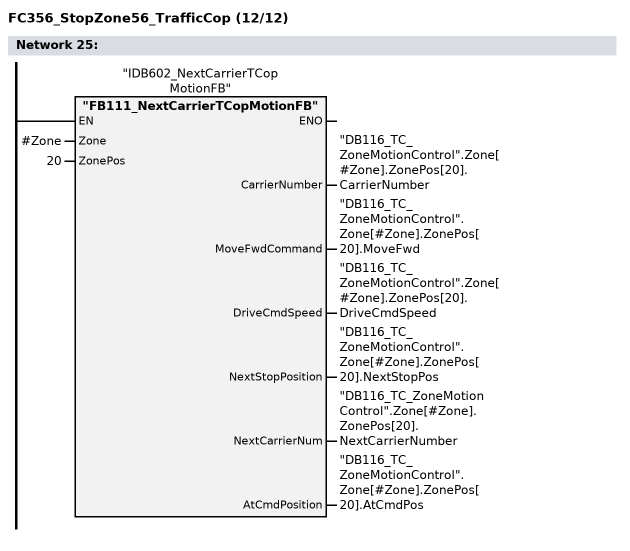
   RUNG wire#powerrail
      "IDB602_NextCarrierTCopMotionFB"(Zone := #Zone, ZonePos := 20, CarrierNumber => "DB116_TC_ZoneMotionControl".Zone[#Zone].ZonePos[20].CarrierNumber, MoveFwdCommand => "DB116_TC_ZoneMotionControl".Zone[#Zone].ZonePos[20].MoveFwd, DriveCmdSpeed => "DB116_TC_ZoneMotionControl".Zone[#Zone].ZonePos[20].DriveCmdSpeed, NextStopPosition => "DB116_TC_ZoneMotionControl".Zone[#Zone].ZonePos[20].NextStopPos, NextCarrierNum => "DB116_TC_ZoneMotionControl".Zone[#Zone].ZonePos[20].NextCarrierNumber, AtCmdPosition => "DB116_TC_ZoneMotionControl".Zone[#Zone].ZonePos[20].AtCmdPos)
   END_RUNG
   // the same network as SCL:
   "IDB602_NextCarrierTCopMotionFB"(Zone := #Zone,   // "FB111_NextCarrierTCopMotionFB"
                           ZonePos := 20,
                           CarrierNumber => "DB116_TC_ZoneMotionControl".Zone[#Zone].ZonePos[20].CarrierNumber,
                           MoveFwdCommand => "DB116_TC_ZoneMotionControl".Zone[#Zone].ZonePos[20].MoveFwd,
                           DriveCmdSpeed => "DB116_TC_ZoneMotionControl".Zone[#Zone].ZonePos[20].DriveCmdSpeed,
                           NextStopPosition => "DB116_TC_ZoneMotionControl".Zone[#Zone].ZonePos[20].NextStopPos,
                           NextCarrierNum => "DB116_TC_ZoneMotionControl".Zone[#Zone].ZonePos[20].NextCarrierNumber,
                           AtCmdPosition => "DB116_TC_ZoneMotionControl".Zone[#Zone].ZonePos[20].AtCmdPos);
END_REGION
END_FUNCTION

FUNCTION "FC357_StopZone57_TrafficCop" : Void   // FC357, LAD
{ S7_Optimized_Access := 'FALSE' }
VERSION : 0.1
   VAR_INPUT
      Zone : Int;
   END_VAR
   VAR_TEMP
      TrafficCopCarrier : Int;
      CarrierMotionZn : Array[0..40] of "UDT_ZoneCarrierStatus";
   END_VAR
BEGIN

REGION Network 1
   // **********************************************************************************************************************
   // 
   // Zone Function Block.  Static setup of all Zone Parameters.  Traffic Cop Setup Logic - Handles all motion and carrier movement logic based on interdependence of Each Carrier in Zone # Passed from Main program Call in OB1 
   // 
   // **********************************************************************************************************************
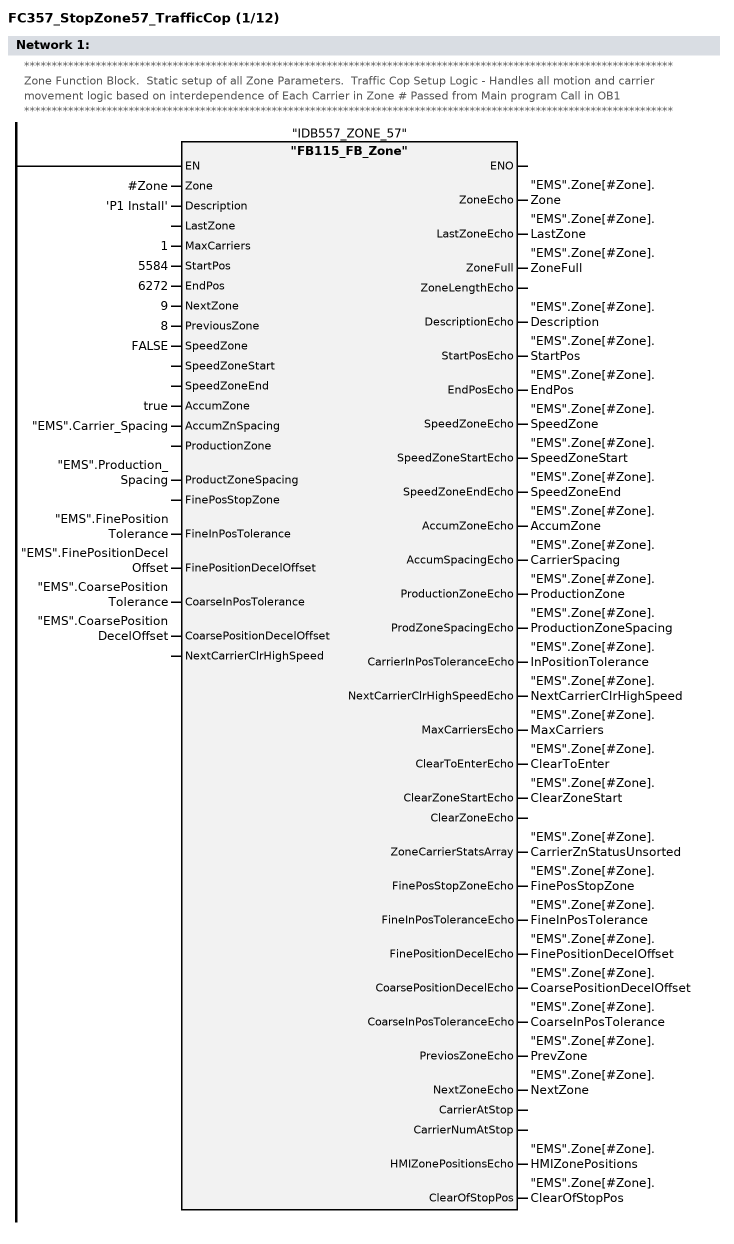
   RUNG wire#powerrail
      "IDB557_ZONE_57"(Zone := #Zone, Description := 'P1 Install', LastZone :=, MaxCarriers := 1, StartPos := 5584, EndPos := 6272, NextZone := 9, PreviousZone := 8, SpeedZone := FALSE, SpeedZoneStart :=, SpeedZoneEnd :=, AccumZone := true, AccumZnSpacing := "EMS".Carrier_Spacing, ProductionZone :=, ProductZoneSpacing := "EMS".Production_Spacing, FinePosStopZone :=, FineInPosTolerance := "EMS".FinePositionTolerance, FinePositionDecelOffset := "EMS".FinePositionDecelOffset, CoarseInPosTolerance := "EMS".CoarsePositionTolerance, CoarsePositionDecelOffset := "EMS".CoarsePositionDecelOffset, NextCarrierClrHighSpeed :=, ZoneEcho => "EMS".Zone[#Zone].Zone, LastZoneEcho => "EMS".Zone[#Zone].LastZone, ZoneFull => "EMS".Zone[#Zone].ZoneFull, ZoneLengthEcho =>, DescriptionEcho => "EMS".Zone[#Zone].Description, StartPosEcho => "EMS".Zone[#Zone].StartPos, EndPosEcho => "EMS".Zone[#Zone].EndPos, SpeedZoneEcho => "EMS".Zone[#Zone].SpeedZone, SpeedZoneStartEcho => "EMS".Zone[#Zone].SpeedZoneStart, SpeedZoneEndEcho => "EMS".Zone[#Zone].SpeedZoneEnd, AccumZoneEcho => "EMS".Zone[#Zone].AccumZone, AccumSpacingEcho => "EMS".Zone[#Zone].CarrierSpacing, ProductionZoneEcho => "EMS".Zone[#Zone].ProductionZone, ProdZoneSpacingEcho => "EMS".Zone[#Zone].ProductionZoneSpacing, CarrierInPosToleranceEcho => "EMS".Zone[#Zone].InPositionTolerance, NextCarrierClrHighSpeedEcho => "EMS".Zone[#Zone].NextCarrierClrHighSpeed, MaxCarriersEcho => "EMS".Zone[#Zone].MaxCarriers, ClearToEnterEcho => "EMS".Zone[#Zone].ClearToEnter, ClearZoneStartEcho => "EMS".Zone[#Zone].ClearZoneStart, ClearZoneEcho =>, ZoneCarrierStatsArray => "EMS".Zone[#Zone].CarrierZnStatusUnsorted, FinePosStopZoneEcho => "EMS".Zone[#Zone].FinePosStopZone, FineInPosToleranceEcho => "EMS".Zone[#Zone].FineInPosTolerance, FinePositionDecelEcho => "EMS".Zone[#Zone].FinePositionDecelOffset, CoarsePositionDecelEcho => "EMS".Zone[#Zone].CoarsePositionDecelOffset, CoarseInPosToleranceEcho => "EMS".Zone[#Zone].CoarseInPosTolerance, PreviosZoneEcho => "EMS".Zone[#Zone].PrevZone, NextZoneEcho => "EMS".Zone[#Zone].NextZone, CarrierAtStop =>, CarrierNumAtStop =>, HMIZonePositionsEcho => "EMS".Zone[#Zone].HMIZonePositions, ClearOfStopPos => "EMS".Zone[#Zone].ClearOfStopPos)
   END_RUNG
   // the same network as SCL:
   "IDB557_ZONE_57"(Zone := #Zone,   // "FB115_FB_Zone"
                    Description := 'P1 Install',
                    MaxCarriers := 1,
                    StartPos := 5584,
                    EndPos := 6272,
                    NextZone := 9,
                    PreviousZone := 8,
                    SpeedZone := FALSE,
                    AccumZone := true,
                    AccumZnSpacing := "EMS".Carrier_Spacing,
                    ProductZoneSpacing := "EMS".Production_Spacing,
                    FineInPosTolerance := "EMS".FinePositionTolerance,
                    FinePositionDecelOffset := "EMS".FinePositionDecelOffset,
                    CoarseInPosTolerance := "EMS".CoarsePositionTolerance,
                    CoarsePositionDecelOffset := "EMS".CoarsePositionDecelOffset,
                    ZoneEcho => "EMS".Zone[#Zone].Zone,
                    LastZoneEcho => "EMS".Zone[#Zone].LastZone,
                    ZoneFull => "EMS".Zone[#Zone].ZoneFull,
                    DescriptionEcho => "EMS".Zone[#Zone].Description,
                    StartPosEcho => "EMS".Zone[#Zone].StartPos,
                    EndPosEcho => "EMS".Zone[#Zone].EndPos,
                    SpeedZoneEcho => "EMS".Zone[#Zone].SpeedZone,
                    SpeedZoneStartEcho => "EMS".Zone[#Zone].SpeedZoneStart,
                    SpeedZoneEndEcho => "EMS".Zone[#Zone].SpeedZoneEnd,
                    AccumZoneEcho => "EMS".Zone[#Zone].AccumZone,
                    AccumSpacingEcho => "EMS".Zone[#Zone].CarrierSpacing,
                    ProductionZoneEcho => "EMS".Zone[#Zone].ProductionZone,
                    ProdZoneSpacingEcho => "EMS".Zone[#Zone].ProductionZoneSpacing,
                    CarrierInPosToleranceEcho => "EMS".Zone[#Zone].InPositionTolerance,
                    NextCarrierClrHighSpeedEcho => "EMS".Zone[#Zone].NextCarrierClrHighSpeed,
                    MaxCarriersEcho => "EMS".Zone[#Zone].MaxCarriers,
                    ClearToEnterEcho => "EMS".Zone[#Zone].ClearToEnter,
                    ClearZoneStartEcho => "EMS".Zone[#Zone].ClearZoneStart,
                    ZoneCarrierStatsArray => "EMS".Zone[#Zone].CarrierZnStatusUnsorted,
                    FinePosStopZoneEcho => "EMS".Zone[#Zone].FinePosStopZone,
                    FineInPosToleranceEcho => "EMS".Zone[#Zone].FineInPosTolerance,
                    FinePositionDecelEcho => "EMS".Zone[#Zone].FinePositionDecelOffset,
                    CoarsePositionDecelEcho => "EMS".Zone[#Zone].CoarsePositionDecelOffset,
                    CoarseInPosToleranceEcho => "EMS".Zone[#Zone].CoarseInPosTolerance,
                    PreviosZoneEcho => "EMS".Zone[#Zone].PrevZone,
                    NextZoneEcho => "EMS".Zone[#Zone].NextZone,
                    HMIZonePositionsEcho => "EMS".Zone[#Zone].HMIZonePositions,
                    ClearOfStopPos => "EMS".Zone[#Zone].ClearOfStopPos);
END_REGION

REGION Network 2
   // *********************************************************************************************************************
   // Carrier Sort Function FC202 - Sorts Carriers in Called Zone to place in correct sequence within  zone. Zones are divided into position based on MaxCarriers allowed in zone as set in the zone setup function block. 
   // 
   // **********************************************************************************************************************
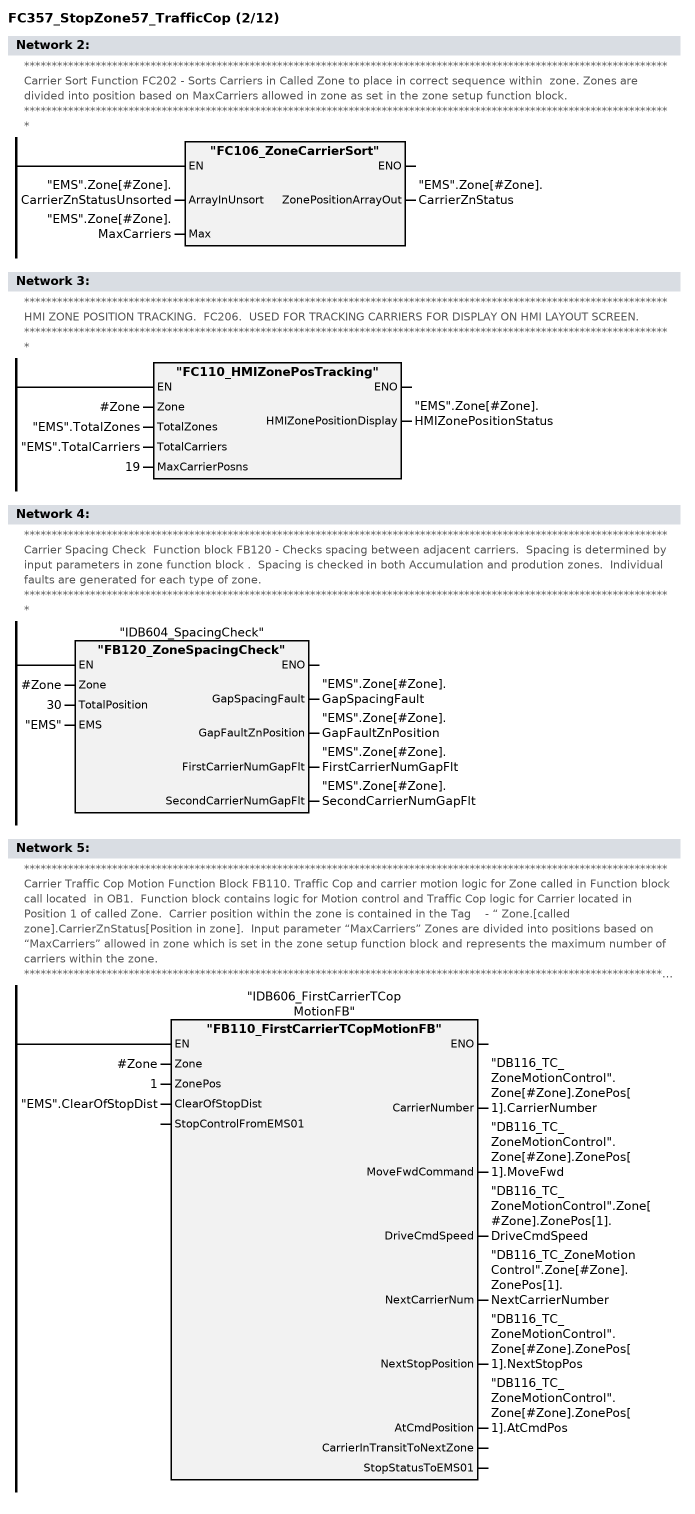
   RUNG wire#powerrail
      "FC106_ZoneCarrierSort"(ArrayInUnsort := "EMS".Zone[#Zone].CarrierZnStatusUnsorted, Max := "EMS".Zone[#Zone].MaxCarriers, ZonePositionArrayOut => "EMS".Zone[#Zone].CarrierZnStatus)
   END_RUNG
   // the same network as SCL:
   "FC106_ZoneCarrierSort"(ArrayInUnsort := "EMS".Zone[#Zone].CarrierZnStatusUnsorted,
                           Max := "EMS".Zone[#Zone].MaxCarriers,
                           ZonePositionArrayOut => "EMS".Zone[#Zone].CarrierZnStatus);
END_REGION

REGION Network 3
   // *********************************************************************************************************************
   // HMI ZONE POSITION TRACKING.  FC206.  USED FOR TRACKING CARRIERS FOR DISPLAY ON HMI LAYOUT SCREEN. 
   // **********************************************************************************************************************
   RUNG wire#powerrail
      "FC110_HMIZonePosTracking"(Zone := #Zone, TotalZones := "EMS".TotalZones, TotalCarriers := "EMS".TotalCarriers, MaxCarrierPosns := 19, HMIZonePositionDisplay => "EMS".Zone[#Zone].HMIZonePositionStatus)
   END_RUNG
   // the same network as SCL:
   "FC110_HMIZonePosTracking"(Zone := #Zone,
                           TotalZones := "EMS".TotalZones,
                           TotalCarriers := "EMS".TotalCarriers,
                           MaxCarrierPosns := 19,
                           HMIZonePositionDisplay => "EMS".Zone[#Zone].HMIZonePositionStatus);
END_REGION

REGION Network 4
   // *********************************************************************************************************************
   // 
   // Carrier Spacing Check  Function block FB120 - Checks spacing between adjacent carriers.  Spacing is determined by input parameters in zone function block .  Spacing is checked in both Accumulation and prodution zones.  Individual faults are generated for each type of zone.
   // 
   // **********************************************************************************************************************
   RUNG wire#powerrail
      "IDB604_SpacingCheck"(Zone := #Zone, TotalPosition := 30, EMS := "EMS", GapSpacingFault => "EMS".Zone[#Zone].GapSpacingFault, GapFaultZnPosition => "EMS".Zone[#Zone].GapFaultZnPosition, FirstCarrierNumGapFlt => "EMS".Zone[#Zone].FirstCarrierNumGapFlt, SecondCarrierNumGapFlt => "EMS".Zone[#Zone].SecondCarrierNumGapFlt)
   END_RUNG
   // the same network as SCL:
   "IDB604_SpacingCheck"(Zone := #Zone,   // "FB120_ZoneSpacingCheck"
                         TotalPosition := 30,
                         EMS := "EMS",
                         GapSpacingFault => "EMS".Zone[#Zone].GapSpacingFault,
                         GapFaultZnPosition => "EMS".Zone[#Zone].GapFaultZnPosition,
                         FirstCarrierNumGapFlt => "EMS".Zone[#Zone].FirstCarrierNumGapFlt,
                         SecondCarrierNumGapFlt => "EMS".Zone[#Zone].SecondCarrierNumGapFlt);
END_REGION

REGION Network 5
   // *********************************************************************************************************************
   // 
   // Carrier Traffic Cop Motion Function Block FB110. Traffic Cop and carrier motion logic for Zone called in Function block call located  in OB1.  Function block contains logic for Motion control and Traffic Cop logic for Carrier located in Position 1 of called Zone.  Carrier position within the zone is contained in the Tag    - “ Zone.[called zone].CarrierZnStatus[Position in zone].  Input parameter “MaxCarriers” Zones are divided into positions based on “MaxCarriers” allowed in zone which is set in the zone setup function block and represents the maximum number of carriers within the zone. 
   // 
   // **********************************************************************************************************************
   RUNG wire#powerrail
      "IDB606_FirstCarrierTCopMotionFB"(Zone := #Zone, ZonePos := 1, ClearOfStopDist := "EMS".ClearOfStopDist, CarrierNumber => "DB116_TC_ZoneMotionControl".Zone[#Zone].ZonePos[1].CarrierNumber, MoveFwdCommand => "DB116_TC_ZoneMotionControl".Zone[#Zone].ZonePos[1].MoveFwd, DriveCmdSpeed => "DB116_TC_ZoneMotionControl".Zone[#Zone].ZonePos[1].DriveCmdSpeed, NextCarrierNum => "DB116_TC_ZoneMotionControl".Zone[#Zone].ZonePos[1].NextCarrierNumber, NextStopPosition => "DB116_TC_ZoneMotionControl".Zone[#Zone].ZonePos[1].NextStopPos, AtCmdPosition => "DB116_TC_ZoneMotionControl".Zone[#Zone].ZonePos[1].AtCmdPos, CarrierInTransitToNextZone =>, StopControlFromEMS01 :=, StopStatusToEMS01 =>)
   END_RUNG
   // the same network as SCL:
   "IDB606_FirstCarrierTCopMotionFB"(Zone := #Zone,   // "FB110_FirstCarrierTCopMotionFB"
                           ZonePos := 1,
                           ClearOfStopDist := "EMS".ClearOfStopDist,
                           CarrierNumber => "DB116_TC_ZoneMotionControl".Zone[#Zone].ZonePos[1].CarrierNumber,
                           MoveFwdCommand => "DB116_TC_ZoneMotionControl".Zone[#Zone].ZonePos[1].MoveFwd,
                           DriveCmdSpeed => "DB116_TC_ZoneMotionControl".Zone[#Zone].ZonePos[1].DriveCmdSpeed,
                           NextCarrierNum => "DB116_TC_ZoneMotionControl".Zone[#Zone].ZonePos[1].NextCarrierNumber,
                           NextStopPosition => "DB116_TC_ZoneMotionControl".Zone[#Zone].ZonePos[1].NextStopPos,
                           AtCmdPosition => "DB116_TC_ZoneMotionControl".Zone[#Zone].ZonePos[1].AtCmdPos);
END_REGION

REGION Network 6
   // *********************************************************************************************************************
   // 
   // Carrier Traffic Cop Motion Function Block FB111. Traffic Cop and carrier motion logic for Zone called in Function block call located  in OB1.  Function block contains logic for Motion control and Traffic Cop logic for Carrier located in Position 2 of called Zone.  Carrier position within the zone is contained in the Tag    - “ Zone.[called zone].CarrierZnStatus[Position in zone].  Input parameter “MaxCarriers” Zones are divided into positions based on “MaxCarriers” allowed in zone which is set in the zone setup function block and represents the maximum number of carriers within the zone. 
   // 
   // **********************************************************************************************************************
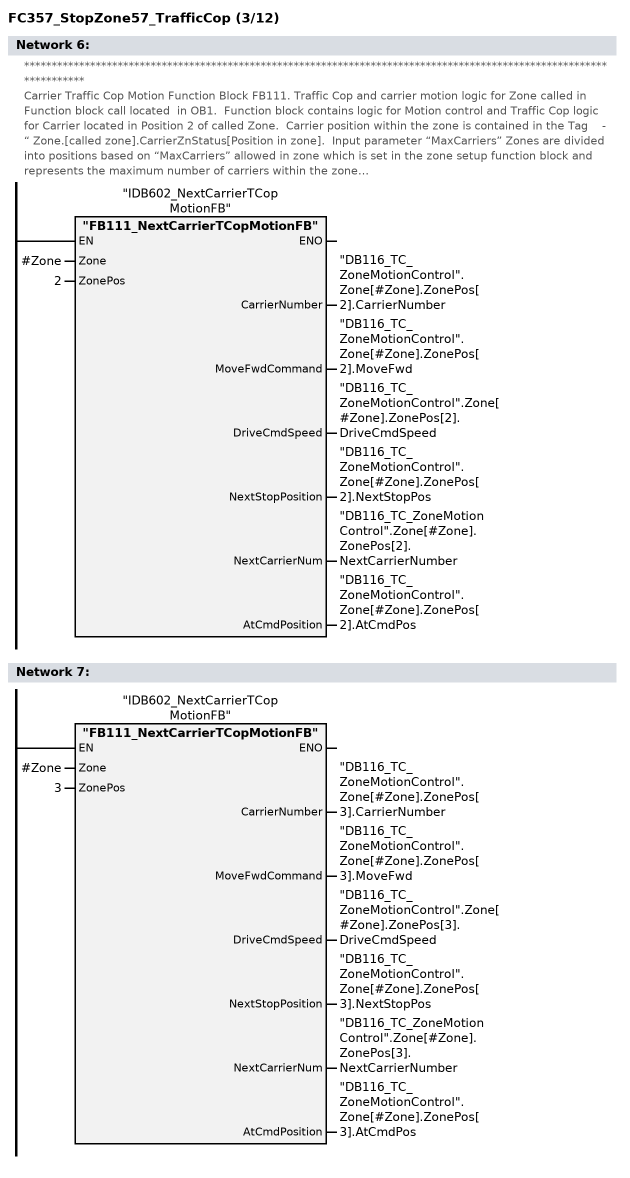
   RUNG wire#powerrail
      "IDB602_NextCarrierTCopMotionFB"(Zone := #Zone, ZonePos := 2, CarrierNumber => "DB116_TC_ZoneMotionControl".Zone[#Zone].ZonePos[2].CarrierNumber, MoveFwdCommand => "DB116_TC_ZoneMotionControl".Zone[#Zone].ZonePos[2].MoveFwd, DriveCmdSpeed => "DB116_TC_ZoneMotionControl".Zone[#Zone].ZonePos[2].DriveCmdSpeed, NextStopPosition => "DB116_TC_ZoneMotionControl".Zone[#Zone].ZonePos[2].NextStopPos, NextCarrierNum => "DB116_TC_ZoneMotionControl".Zone[#Zone].ZonePos[2].NextCarrierNumber, AtCmdPosition => "DB116_TC_ZoneMotionControl".Zone[#Zone].ZonePos[2].AtCmdPos)
   END_RUNG
   // the same network as SCL:
   "IDB602_NextCarrierTCopMotionFB"(Zone := #Zone,   // "FB111_NextCarrierTCopMotionFB"
                           ZonePos := 2,
                           CarrierNumber => "DB116_TC_ZoneMotionControl".Zone[#Zone].ZonePos[2].CarrierNumber,
                           MoveFwdCommand => "DB116_TC_ZoneMotionControl".Zone[#Zone].ZonePos[2].MoveFwd,
                           DriveCmdSpeed => "DB116_TC_ZoneMotionControl".Zone[#Zone].ZonePos[2].DriveCmdSpeed,
                           NextStopPosition => "DB116_TC_ZoneMotionControl".Zone[#Zone].ZonePos[2].NextStopPos,
                           NextCarrierNum => "DB116_TC_ZoneMotionControl".Zone[#Zone].ZonePos[2].NextCarrierNumber,
                           AtCmdPosition => "DB116_TC_ZoneMotionControl".Zone[#Zone].ZonePos[2].AtCmdPos);
END_REGION

REGION Network 7
   RUNG wire#powerrail
      "IDB602_NextCarrierTCopMotionFB"(Zone := #Zone, ZonePos := 3, CarrierNumber => "DB116_TC_ZoneMotionControl".Zone[#Zone].ZonePos[3].CarrierNumber, MoveFwdCommand => "DB116_TC_ZoneMotionControl".Zone[#Zone].ZonePos[3].MoveFwd, DriveCmdSpeed => "DB116_TC_ZoneMotionControl".Zone[#Zone].ZonePos[3].DriveCmdSpeed, NextStopPosition => "DB116_TC_ZoneMotionControl".Zone[#Zone].ZonePos[3].NextStopPos, NextCarrierNum => "DB116_TC_ZoneMotionControl".Zone[#Zone].ZonePos[3].NextCarrierNumber, AtCmdPosition => "DB116_TC_ZoneMotionControl".Zone[#Zone].ZonePos[3].AtCmdPos)
   END_RUNG
   // the same network as SCL:
   "IDB602_NextCarrierTCopMotionFB"(Zone := #Zone,   // "FB111_NextCarrierTCopMotionFB"
                           ZonePos := 3,
                           CarrierNumber => "DB116_TC_ZoneMotionControl".Zone[#Zone].ZonePos[3].CarrierNumber,
                           MoveFwdCommand => "DB116_TC_ZoneMotionControl".Zone[#Zone].ZonePos[3].MoveFwd,
                           DriveCmdSpeed => "DB116_TC_ZoneMotionControl".Zone[#Zone].ZonePos[3].DriveCmdSpeed,
                           NextStopPosition => "DB116_TC_ZoneMotionControl".Zone[#Zone].ZonePos[3].NextStopPos,
                           NextCarrierNum => "DB116_TC_ZoneMotionControl".Zone[#Zone].ZonePos[3].NextCarrierNumber,
                           AtCmdPosition => "DB116_TC_ZoneMotionControl".Zone[#Zone].ZonePos[3].AtCmdPos);
END_REGION

REGION Network 8
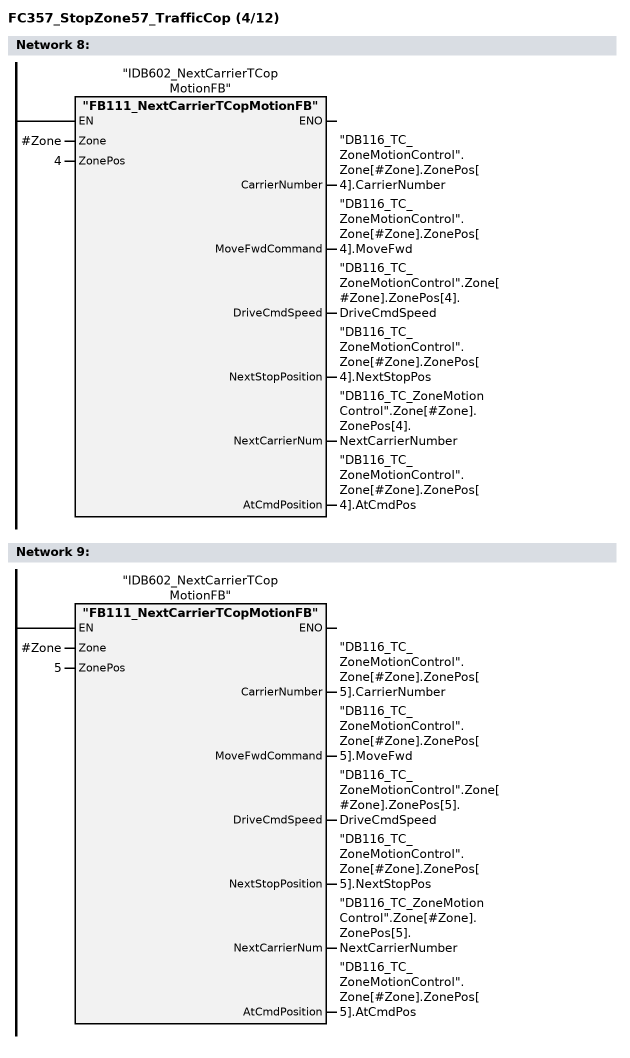
   RUNG wire#powerrail
      "IDB602_NextCarrierTCopMotionFB"(Zone := #Zone, ZonePos := 4, CarrierNumber => "DB116_TC_ZoneMotionControl".Zone[#Zone].ZonePos[4].CarrierNumber, MoveFwdCommand => "DB116_TC_ZoneMotionControl".Zone[#Zone].ZonePos[4].MoveFwd, DriveCmdSpeed => "DB116_TC_ZoneMotionControl".Zone[#Zone].ZonePos[4].DriveCmdSpeed, NextStopPosition => "DB116_TC_ZoneMotionControl".Zone[#Zone].ZonePos[4].NextStopPos, NextCarrierNum => "DB116_TC_ZoneMotionControl".Zone[#Zone].ZonePos[4].NextCarrierNumber, AtCmdPosition => "DB116_TC_ZoneMotionControl".Zone[#Zone].ZonePos[4].AtCmdPos)
   END_RUNG
   // the same network as SCL:
   "IDB602_NextCarrierTCopMotionFB"(Zone := #Zone,   // "FB111_NextCarrierTCopMotionFB"
                           ZonePos := 4,
                           CarrierNumber => "DB116_TC_ZoneMotionControl".Zone[#Zone].ZonePos[4].CarrierNumber,
                           MoveFwdCommand => "DB116_TC_ZoneMotionControl".Zone[#Zone].ZonePos[4].MoveFwd,
                           DriveCmdSpeed => "DB116_TC_ZoneMotionControl".Zone[#Zone].ZonePos[4].DriveCmdSpeed,
                           NextStopPosition => "DB116_TC_ZoneMotionControl".Zone[#Zone].ZonePos[4].NextStopPos,
                           NextCarrierNum => "DB116_TC_ZoneMotionControl".Zone[#Zone].ZonePos[4].NextCarrierNumber,
                           AtCmdPosition => "DB116_TC_ZoneMotionControl".Zone[#Zone].ZonePos[4].AtCmdPos);
END_REGION

REGION Network 9
   RUNG wire#powerrail
      "IDB602_NextCarrierTCopMotionFB"(Zone := #Zone, ZonePos := 5, CarrierNumber => "DB116_TC_ZoneMotionControl".Zone[#Zone].ZonePos[5].CarrierNumber, MoveFwdCommand => "DB116_TC_ZoneMotionControl".Zone[#Zone].ZonePos[5].MoveFwd, DriveCmdSpeed => "DB116_TC_ZoneMotionControl".Zone[#Zone].ZonePos[5].DriveCmdSpeed, NextStopPosition => "DB116_TC_ZoneMotionControl".Zone[#Zone].ZonePos[5].NextStopPos, NextCarrierNum => "DB116_TC_ZoneMotionControl".Zone[#Zone].ZonePos[5].NextCarrierNumber, AtCmdPosition => "DB116_TC_ZoneMotionControl".Zone[#Zone].ZonePos[5].AtCmdPos)
   END_RUNG
   // the same network as SCL:
   "IDB602_NextCarrierTCopMotionFB"(Zone := #Zone,   // "FB111_NextCarrierTCopMotionFB"
                           ZonePos := 5,
                           CarrierNumber => "DB116_TC_ZoneMotionControl".Zone[#Zone].ZonePos[5].CarrierNumber,
                           MoveFwdCommand => "DB116_TC_ZoneMotionControl".Zone[#Zone].ZonePos[5].MoveFwd,
                           DriveCmdSpeed => "DB116_TC_ZoneMotionControl".Zone[#Zone].ZonePos[5].DriveCmdSpeed,
                           NextStopPosition => "DB116_TC_ZoneMotionControl".Zone[#Zone].ZonePos[5].NextStopPos,
                           NextCarrierNum => "DB116_TC_ZoneMotionControl".Zone[#Zone].ZonePos[5].NextCarrierNumber,
                           AtCmdPosition => "DB116_TC_ZoneMotionControl".Zone[#Zone].ZonePos[5].AtCmdPos);
END_REGION

REGION Network 10
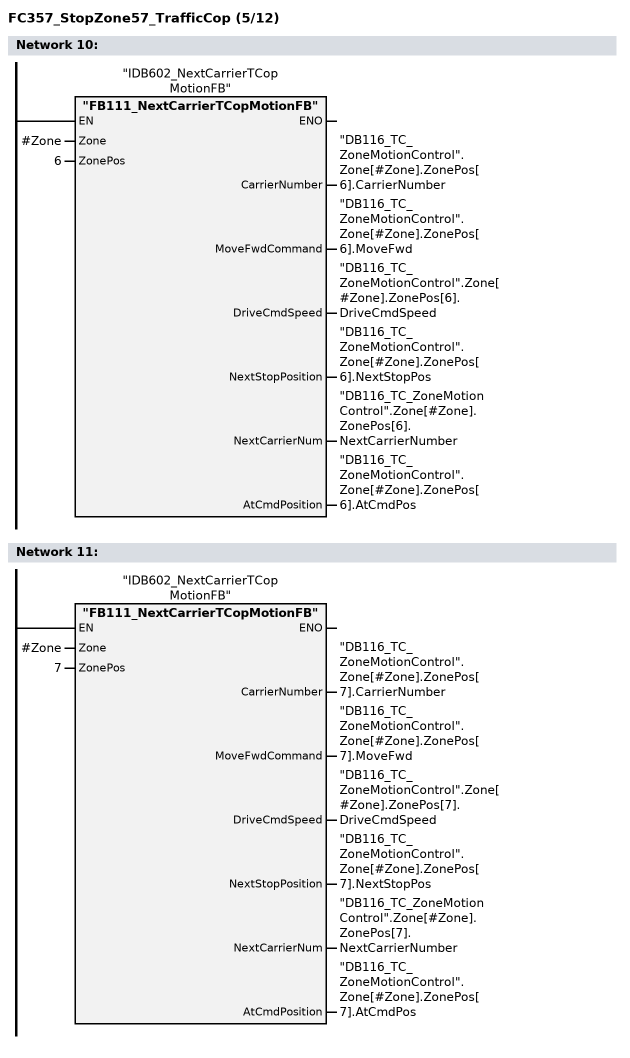
   RUNG wire#powerrail
      "IDB602_NextCarrierTCopMotionFB"(Zone := #Zone, ZonePos := 6, CarrierNumber => "DB116_TC_ZoneMotionControl".Zone[#Zone].ZonePos[6].CarrierNumber, MoveFwdCommand => "DB116_TC_ZoneMotionControl".Zone[#Zone].ZonePos[6].MoveFwd, DriveCmdSpeed => "DB116_TC_ZoneMotionControl".Zone[#Zone].ZonePos[6].DriveCmdSpeed, NextStopPosition => "DB116_TC_ZoneMotionControl".Zone[#Zone].ZonePos[6].NextStopPos, NextCarrierNum => "DB116_TC_ZoneMotionControl".Zone[#Zone].ZonePos[6].NextCarrierNumber, AtCmdPosition => "DB116_TC_ZoneMotionControl".Zone[#Zone].ZonePos[6].AtCmdPos)
   END_RUNG
   // the same network as SCL:
   "IDB602_NextCarrierTCopMotionFB"(Zone := #Zone,   // "FB111_NextCarrierTCopMotionFB"
                           ZonePos := 6,
                           CarrierNumber => "DB116_TC_ZoneMotionControl".Zone[#Zone].ZonePos[6].CarrierNumber,
                           MoveFwdCommand => "DB116_TC_ZoneMotionControl".Zone[#Zone].ZonePos[6].MoveFwd,
                           DriveCmdSpeed => "DB116_TC_ZoneMotionControl".Zone[#Zone].ZonePos[6].DriveCmdSpeed,
                           NextStopPosition => "DB116_TC_ZoneMotionControl".Zone[#Zone].ZonePos[6].NextStopPos,
                           NextCarrierNum => "DB116_TC_ZoneMotionControl".Zone[#Zone].ZonePos[6].NextCarrierNumber,
                           AtCmdPosition => "DB116_TC_ZoneMotionControl".Zone[#Zone].ZonePos[6].AtCmdPos);
END_REGION

REGION Network 11
   RUNG wire#powerrail
      "IDB602_NextCarrierTCopMotionFB"(Zone := #Zone, ZonePos := 7, CarrierNumber => "DB116_TC_ZoneMotionControl".Zone[#Zone].ZonePos[7].CarrierNumber, MoveFwdCommand => "DB116_TC_ZoneMotionControl".Zone[#Zone].ZonePos[7].MoveFwd, DriveCmdSpeed => "DB116_TC_ZoneMotionControl".Zone[#Zone].ZonePos[7].DriveCmdSpeed, NextStopPosition => "DB116_TC_ZoneMotionControl".Zone[#Zone].ZonePos[7].NextStopPos, NextCarrierNum => "DB116_TC_ZoneMotionControl".Zone[#Zone].ZonePos[7].NextCarrierNumber, AtCmdPosition => "DB116_TC_ZoneMotionControl".Zone[#Zone].ZonePos[7].AtCmdPos)
   END_RUNG
   // the same network as SCL:
   "IDB602_NextCarrierTCopMotionFB"(Zone := #Zone,   // "FB111_NextCarrierTCopMotionFB"
                           ZonePos := 7,
                           CarrierNumber => "DB116_TC_ZoneMotionControl".Zone[#Zone].ZonePos[7].CarrierNumber,
                           MoveFwdCommand => "DB116_TC_ZoneMotionControl".Zone[#Zone].ZonePos[7].MoveFwd,
                           DriveCmdSpeed => "DB116_TC_ZoneMotionControl".Zone[#Zone].ZonePos[7].DriveCmdSpeed,
                           NextStopPosition => "DB116_TC_ZoneMotionControl".Zone[#Zone].ZonePos[7].NextStopPos,
                           NextCarrierNum => "DB116_TC_ZoneMotionControl".Zone[#Zone].ZonePos[7].NextCarrierNumber,
                           AtCmdPosition => "DB116_TC_ZoneMotionControl".Zone[#Zone].ZonePos[7].AtCmdPos);
END_REGION

REGION Network 12
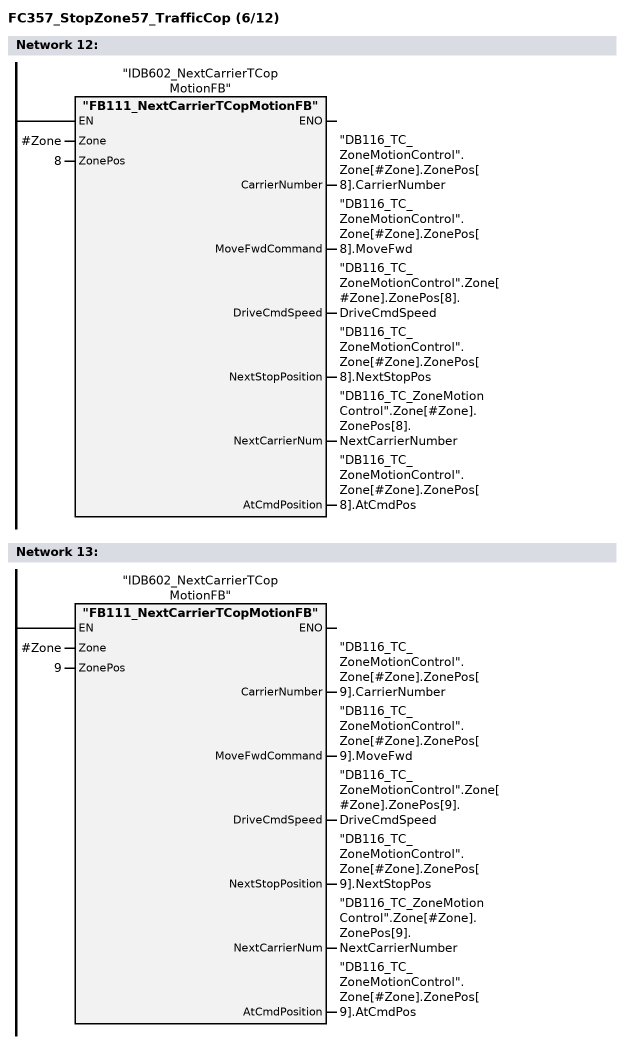
   RUNG wire#powerrail
      "IDB602_NextCarrierTCopMotionFB"(Zone := #Zone, ZonePos := 8, CarrierNumber => "DB116_TC_ZoneMotionControl".Zone[#Zone].ZonePos[8].CarrierNumber, MoveFwdCommand => "DB116_TC_ZoneMotionControl".Zone[#Zone].ZonePos[8].MoveFwd, DriveCmdSpeed => "DB116_TC_ZoneMotionControl".Zone[#Zone].ZonePos[8].DriveCmdSpeed, NextStopPosition => "DB116_TC_ZoneMotionControl".Zone[#Zone].ZonePos[8].NextStopPos, NextCarrierNum => "DB116_TC_ZoneMotionControl".Zone[#Zone].ZonePos[8].NextCarrierNumber, AtCmdPosition => "DB116_TC_ZoneMotionControl".Zone[#Zone].ZonePos[8].AtCmdPos)
   END_RUNG
   // the same network as SCL:
   "IDB602_NextCarrierTCopMotionFB"(Zone := #Zone,   // "FB111_NextCarrierTCopMotionFB"
                           ZonePos := 8,
                           CarrierNumber => "DB116_TC_ZoneMotionControl".Zone[#Zone].ZonePos[8].CarrierNumber,
                           MoveFwdCommand => "DB116_TC_ZoneMotionControl".Zone[#Zone].ZonePos[8].MoveFwd,
                           DriveCmdSpeed => "DB116_TC_ZoneMotionControl".Zone[#Zone].ZonePos[8].DriveCmdSpeed,
                           NextStopPosition => "DB116_TC_ZoneMotionControl".Zone[#Zone].ZonePos[8].NextStopPos,
                           NextCarrierNum => "DB116_TC_ZoneMotionControl".Zone[#Zone].ZonePos[8].NextCarrierNumber,
                           AtCmdPosition => "DB116_TC_ZoneMotionControl".Zone[#Zone].ZonePos[8].AtCmdPos);
END_REGION

REGION Network 13
   RUNG wire#powerrail
      "IDB602_NextCarrierTCopMotionFB"(Zone := #Zone, ZonePos := 9, CarrierNumber => "DB116_TC_ZoneMotionControl".Zone[#Zone].ZonePos[9].CarrierNumber, MoveFwdCommand => "DB116_TC_ZoneMotionControl".Zone[#Zone].ZonePos[9].MoveFwd, DriveCmdSpeed => "DB116_TC_ZoneMotionControl".Zone[#Zone].ZonePos[9].DriveCmdSpeed, NextStopPosition => "DB116_TC_ZoneMotionControl".Zone[#Zone].ZonePos[9].NextStopPos, NextCarrierNum => "DB116_TC_ZoneMotionControl".Zone[#Zone].ZonePos[9].NextCarrierNumber, AtCmdPosition => "DB116_TC_ZoneMotionControl".Zone[#Zone].ZonePos[9].AtCmdPos)
   END_RUNG
   // the same network as SCL:
   "IDB602_NextCarrierTCopMotionFB"(Zone := #Zone,   // "FB111_NextCarrierTCopMotionFB"
                           ZonePos := 9,
                           CarrierNumber => "DB116_TC_ZoneMotionControl".Zone[#Zone].ZonePos[9].CarrierNumber,
                           MoveFwdCommand => "DB116_TC_ZoneMotionControl".Zone[#Zone].ZonePos[9].MoveFwd,
                           DriveCmdSpeed => "DB116_TC_ZoneMotionControl".Zone[#Zone].ZonePos[9].DriveCmdSpeed,
                           NextStopPosition => "DB116_TC_ZoneMotionControl".Zone[#Zone].ZonePos[9].NextStopPos,
                           NextCarrierNum => "DB116_TC_ZoneMotionControl".Zone[#Zone].ZonePos[9].NextCarrierNumber,
                           AtCmdPosition => "DB116_TC_ZoneMotionControl".Zone[#Zone].ZonePos[9].AtCmdPos);
END_REGION

REGION Network 14
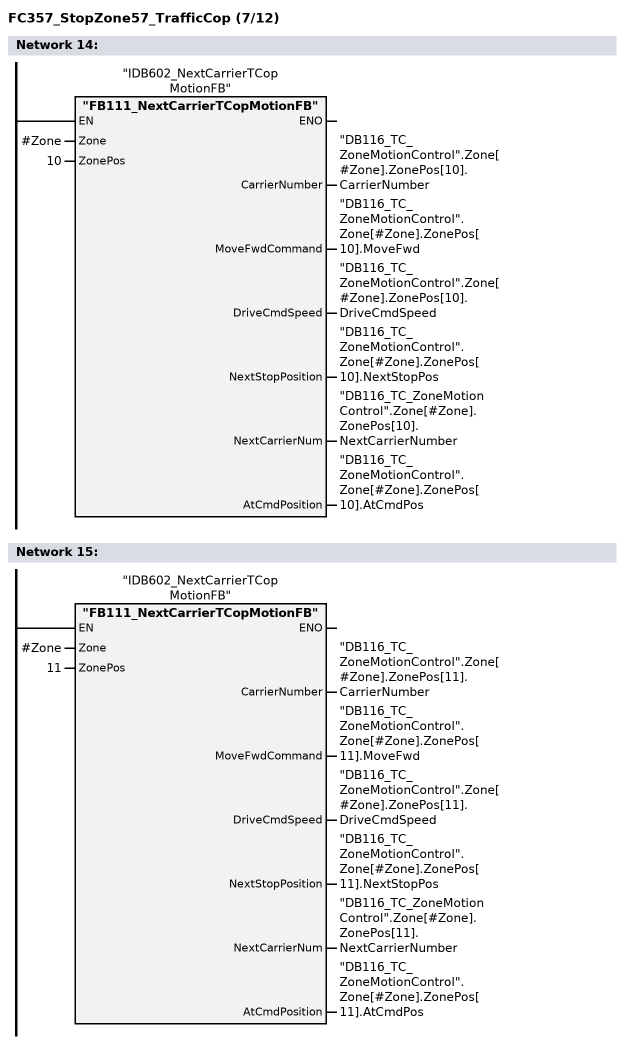
   RUNG wire#powerrail
      "IDB602_NextCarrierTCopMotionFB"(Zone := #Zone, ZonePos := 10, CarrierNumber => "DB116_TC_ZoneMotionControl".Zone[#Zone].ZonePos[10].CarrierNumber, MoveFwdCommand => "DB116_TC_ZoneMotionControl".Zone[#Zone].ZonePos[10].MoveFwd, DriveCmdSpeed => "DB116_TC_ZoneMotionControl".Zone[#Zone].ZonePos[10].DriveCmdSpeed, NextStopPosition => "DB116_TC_ZoneMotionControl".Zone[#Zone].ZonePos[10].NextStopPos, NextCarrierNum => "DB116_TC_ZoneMotionControl".Zone[#Zone].ZonePos[10].NextCarrierNumber, AtCmdPosition => "DB116_TC_ZoneMotionControl".Zone[#Zone].ZonePos[10].AtCmdPos)
   END_RUNG
   // the same network as SCL:
   "IDB602_NextCarrierTCopMotionFB"(Zone := #Zone,   // "FB111_NextCarrierTCopMotionFB"
                           ZonePos := 10,
                           CarrierNumber => "DB116_TC_ZoneMotionControl".Zone[#Zone].ZonePos[10].CarrierNumber,
                           MoveFwdCommand => "DB116_TC_ZoneMotionControl".Zone[#Zone].ZonePos[10].MoveFwd,
                           DriveCmdSpeed => "DB116_TC_ZoneMotionControl".Zone[#Zone].ZonePos[10].DriveCmdSpeed,
                           NextStopPosition => "DB116_TC_ZoneMotionControl".Zone[#Zone].ZonePos[10].NextStopPos,
                           NextCarrierNum => "DB116_TC_ZoneMotionControl".Zone[#Zone].ZonePos[10].NextCarrierNumber,
                           AtCmdPosition => "DB116_TC_ZoneMotionControl".Zone[#Zone].ZonePos[10].AtCmdPos);
END_REGION

REGION Network 15
   RUNG wire#powerrail
      "IDB602_NextCarrierTCopMotionFB"(Zone := #Zone, ZonePos := 11, CarrierNumber => "DB116_TC_ZoneMotionControl".Zone[#Zone].ZonePos[11].CarrierNumber, MoveFwdCommand => "DB116_TC_ZoneMotionControl".Zone[#Zone].ZonePos[11].MoveFwd, DriveCmdSpeed => "DB116_TC_ZoneMotionControl".Zone[#Zone].ZonePos[11].DriveCmdSpeed, NextStopPosition => "DB116_TC_ZoneMotionControl".Zone[#Zone].ZonePos[11].NextStopPos, NextCarrierNum => "DB116_TC_ZoneMotionControl".Zone[#Zone].ZonePos[11].NextCarrierNumber, AtCmdPosition => "DB116_TC_ZoneMotionControl".Zone[#Zone].ZonePos[11].AtCmdPos)
   END_RUNG
   // the same network as SCL:
   "IDB602_NextCarrierTCopMotionFB"(Zone := #Zone,   // "FB111_NextCarrierTCopMotionFB"
                           ZonePos := 11,
                           CarrierNumber => "DB116_TC_ZoneMotionControl".Zone[#Zone].ZonePos[11].CarrierNumber,
                           MoveFwdCommand => "DB116_TC_ZoneMotionControl".Zone[#Zone].ZonePos[11].MoveFwd,
                           DriveCmdSpeed => "DB116_TC_ZoneMotionControl".Zone[#Zone].ZonePos[11].DriveCmdSpeed,
                           NextStopPosition => "DB116_TC_ZoneMotionControl".Zone[#Zone].ZonePos[11].NextStopPos,
                           NextCarrierNum => "DB116_TC_ZoneMotionControl".Zone[#Zone].ZonePos[11].NextCarrierNumber,
                           AtCmdPosition => "DB116_TC_ZoneMotionControl".Zone[#Zone].ZonePos[11].AtCmdPos);
END_REGION

REGION Network 16
